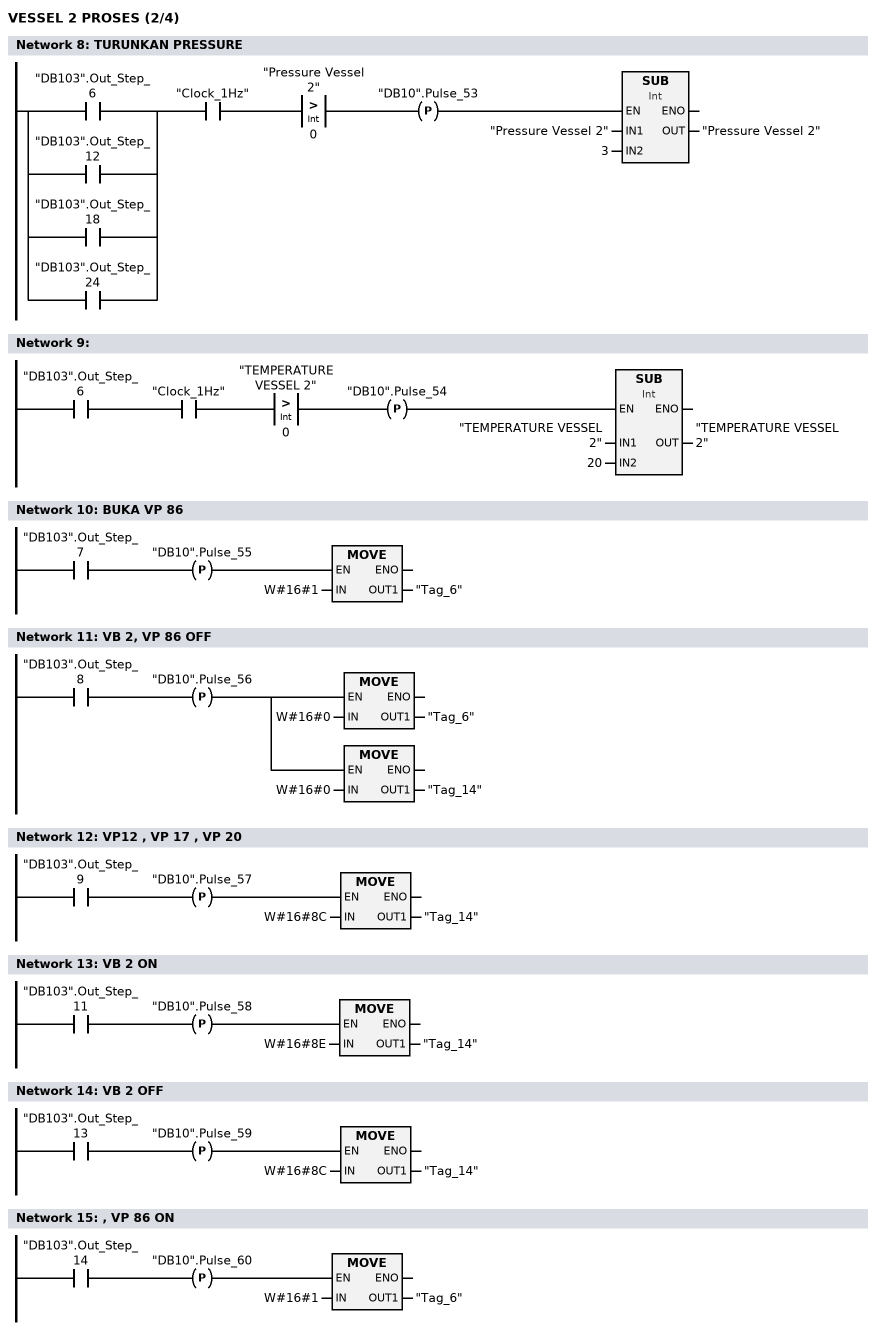
   RUNG wire#powerrail
      Contact( "DB103".Out_Step_6 )
      wire#w1
      Contact( "Clock_1Hz" )
      { S7_Templates := "SrcType := Int" } GT_Contact(in1 := "Pressure Vessel 2", in2 := 0)
      P_Trig( "DB10".Pulse_53 )
      { S7_Templates := "SrcType := Int" } Sub(in1 := "Pressure Vessel 2", in2 := 3, out => "Pressure Vessel 2")
   END_RUNG
   RUNG wire#powerrail
      Contact( "DB103".Out_Step_12 )
   END_RUNG wire#w1
   RUNG wire#powerrail
      Contact( "DB103".Out_Step_18 )
   END_RUNG wire#w1
   RUNG wire#powerrail
      Contact( "DB103".Out_Step_24 )
   END_RUNG wire#w1
   // the same network as SCL:
   #_w1 := ("DB103".Out_Step_6 OR "DB103".Out_Step_12 OR "DB103".Out_Step_18 OR "DB103".Out_Step_24) AND "Clock_1Hz" AND ("Pressure Vessel 2" > 0);
   #_w2 := #_w1 AND NOT "DB10".Pulse_53;   // rising edge
   "DB10".Pulse_53 := #_w1;
   IF #_w2 THEN "Pressure Vessel 2" := "Pressure Vessel 2" - 3; END_IF;
END_REGION

REGION Network 9
   RUNG wire#powerrail
      Contact( "DB103".Out_Step_6 )
      Contact( "Clock_1Hz" )
      { S7_Templates := "SrcType := Int" } GT_Contact(in1 := "TEMPERATURE VESSEL 2", in2 := 0)
      P_Trig( "DB10".Pulse_54 )
      { S7_Templates := "SrcType := Int" } Sub(in1 := "TEMPERATURE VESSEL 2", in2 := 20, out => "TEMPERATURE VESSEL 2")
   END_RUNG
   // the same network as SCL:
   #_w1 := "DB103".Out_Step_6 AND "Clock_1Hz" AND ("TEMPERATURE VESSEL 2" > 0);
   #_w2 := #_w1 AND NOT "DB10".Pulse_54;   // rising edge
   "DB10".Pulse_54 := #_w1;
   IF #_w2 THEN "TEMPERATURE VESSEL 2" := "TEMPERATURE VESSEL 2" - 20; END_IF;
END_REGION

REGION Network 10: BUKA VP 86
   RUNG wire#powerrail
      Contact( "DB103".Out_Step_7 )
      P_Trig( "DB10".Pulse_55 )
      Move(in := W#16#1, out1 => "Tag_6")
   END_RUNG
   // the same network as SCL:
   #_w1 := "DB103".Out_Step_7 AND NOT "DB10".Pulse_55;   // rising edge
   "DB10".Pulse_55 := "DB103".Out_Step_7;
   IF #_w1 THEN "Tag_6" := W#16#1; END_IF;
END_REGION

REGION Network 11: VB 2, VP 86 OFF
   RUNG wire#powerrail
      Contact( "DB103".Out_Step_8 )
      P_Trig( "DB10".Pulse_56 )
      wire#w1
      Move(in := W#16#0, out1 => "Tag_6")
   END_RUNG
   RUNG wire#w1
      Move(in := W#16#0, out1 => "Tag_14")
   END_RUNG
   // the same network as SCL:
   #_w1 := "DB103".Out_Step_8 AND NOT "DB10".Pulse_56;   // rising edge
   "DB10".Pulse_56 := "DB103".Out_Step_8;
   IF #_w1 THEN
       "Tag_6" := W#16#0;
       "Tag_14" := W#16#0;
   END_IF;
END_REGION

REGION Network 12: VP12 , VP 17 , VP 20
   RUNG wire#powerrail
      Contact( "DB103".Out_Step_9 )
      P_Trig( "DB10".Pulse_57 )
      Move(in := W#16#8C, out1 => "Tag_14")
   END_RUNG
   // the same network as SCL:
   #_w1 := "DB103".Out_Step_9 AND NOT "DB10".Pulse_57;   // rising edge
   "DB10".Pulse_57 := "DB103".Out_Step_9;
   IF #_w1 THEN "Tag_14" := W#16#8C; END_IF;
END_REGION

REGION Network 13: VB 2 ON
   RUNG wire#powerrail
      Contact( "DB103".Out_Step_11 )
      P_Trig( "DB10".Pulse_58 )
      Move(in := W#16#8E, out1 => "Tag_14")
   END_RUNG
   // the same network as SCL:
   #_w1 := "DB103".Out_Step_11 AND NOT "DB10".Pulse_58;   // rising edge
   "DB10".Pulse_58 := "DB103".Out_Step_11;
   IF #_w1 THEN "Tag_14" := W#16#8E; END_IF;
END_REGION

REGION Network 14: VB 2 OFF
   RUNG wire#powerrail
      Contact( "DB103".Out_Step_13 )
      P_Trig( "DB10".Pulse_59 )
      Move(in := W#16#8C, out1 => "Tag_14")
   END_RUNG
   // the same network as SCL:
   #_w1 := "DB103".Out_Step_13 AND NOT "DB10".Pulse_59;   // rising edge
   "DB10".Pulse_59 := "DB103".Out_Step_13;
   IF #_w1 THEN "Tag_14" := W#16#8C; END_IF;
END_REGION

REGION Network 15: , VP 86 ON
   RUNG wire#powerrail
      Contact( "DB103".Out_Step_14 )
      P_Trig( "DB10".Pulse_60 )
      Move(in := W#16#1, out1 => "Tag_6")
   END_RUNG
   // the same network as SCL:
   #_w1 := "DB103".Out_Step_14 AND NOT "DB10".Pulse_60;   // rising edge
   "DB10".Pulse_60 := "DB103".Out_Step_14;
   IF #_w1 THEN "Tag_6" := W#16#1; END_IF;
END_REGION

REGION Network 16: VP 86 OFF
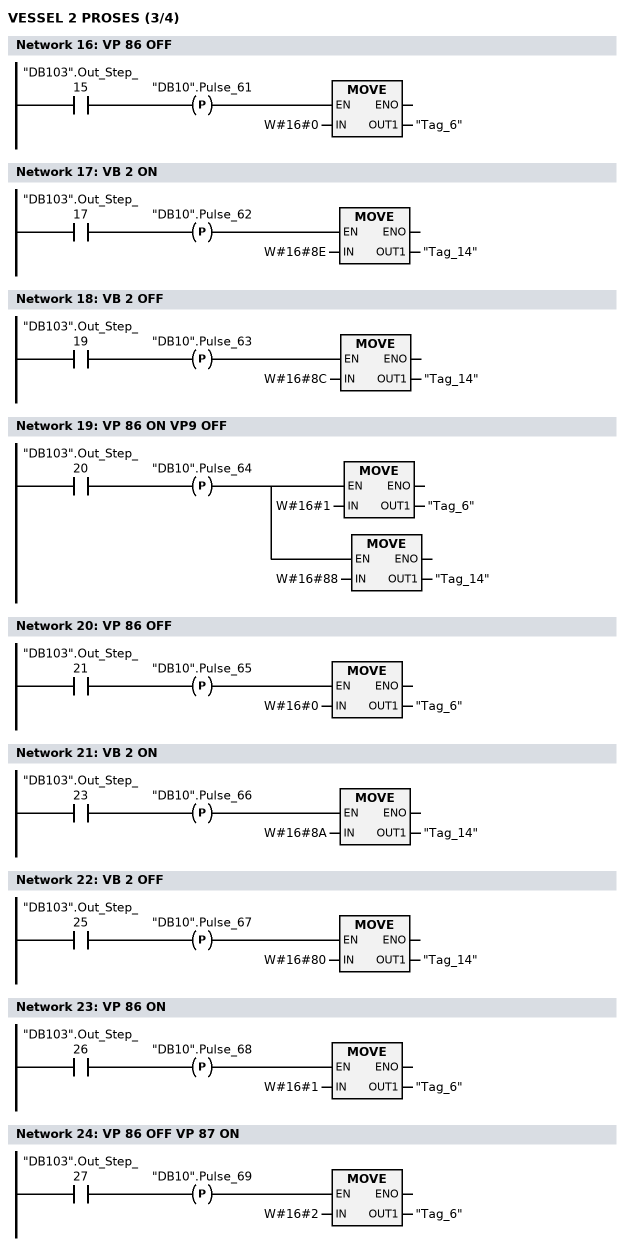
   RUNG wire#powerrail
      Contact( "DB103".Out_Step_15 )
      P_Trig( "DB10".Pulse_61 )
      Move(in := W#16#0, out1 => "Tag_6")
   END_RUNG
   // the same network as SCL:
   #_w1 := "DB103".Out_Step_15 AND NOT "DB10".Pulse_61;   // rising edge
   "DB10".Pulse_61 := "DB103".Out_Step_15;
   IF #_w1 THEN "Tag_6" := W#16#0; END_IF;
END_REGION

REGION Network 17: VB 2 ON
   RUNG wire#powerrail
      Contact( "DB103".Out_Step_17 )
      P_Trig( "DB10".Pulse_62 )
      Move(in := W#16#8E, out1 => "Tag_14")
   END_RUNG
   // the same network as SCL:
   #_w1 := "DB103".Out_Step_17 AND NOT "DB10".Pulse_62;   // rising edge
   "DB10".Pulse_62 := "DB103".Out_Step_17;
   IF #_w1 THEN "Tag_14" := W#16#8E; END_IF;
END_REGION

REGION Network 18: VB 2 OFF
   RUNG wire#powerrail
      Contact( "DB103".Out_Step_19 )
      P_Trig( "DB10".Pulse_63 )
      Move(in := W#16#8C, out1 => "Tag_14")
   END_RUNG
   // the same network as SCL:
   #_w1 := "DB103".Out_Step_19 AND NOT "DB10".Pulse_63;   // rising edge
   "DB10".Pulse_63 := "DB103".Out_Step_19;
   IF #_w1 THEN "Tag_14" := W#16#8C; END_IF;
END_REGION

REGION Network 19: VP 86 ON VP9 OFF
   RUNG wire#powerrail
      Contact( "DB103".Out_Step_20 )
      P_Trig( "DB10".Pulse_64 )
      wire#w1
      Move(in := W#16#1, out1 => "Tag_6")
   END_RUNG
   RUNG wire#w1
      Move(in := W#16#88, out1 => "Tag_14")
   END_RUNG
   // the same network as SCL:
   #_w1 := "DB103".Out_Step_20 AND NOT "DB10".Pulse_64;   // rising edge
   "DB10".Pulse_64 := "DB103".Out_Step_20;
   IF #_w1 THEN
       "Tag_6" := W#16#1;
       "Tag_14" := W#16#88;
   END_IF;
END_REGION

REGION Network 20: VP 86 OFF
   RUNG wire#powerrail
      Contact( "DB103".Out_Step_21 )
      P_Trig( "DB10".Pulse_65 )
      Move(in := W#16#0, out1 => "Tag_6")
   END_RUNG
   // the same network as SCL:
   #_w1 := "DB103".Out_Step_21 AND NOT "DB10".Pulse_65;   // rising edge
   "DB10".Pulse_65 := "DB103".Out_Step_21;
   IF #_w1 THEN "Tag_6" := W#16#0; END_IF;
END_REGION

REGION Network 21: VB 2 ON
   RUNG wire#powerrail
      Contact( "DB103".Out_Step_23 )
      P_Trig( "DB10".Pulse_66 )
      Move(in := W#16#8A, out1 => "Tag_14")
   END_RUNG
   // the same network as SCL:
   #_w1 := "DB103".Out_Step_23 AND NOT "DB10".Pulse_66;   // rising edge
   "DB10".Pulse_66 := "DB103".Out_Step_23;
   IF #_w1 THEN "Tag_14" := W#16#8A; END_IF;
END_REGION

REGION Network 22: VB 2 OFF
   RUNG wire#powerrail
      Contact( "DB103".Out_Step_25 )
      P_Trig( "DB10".Pulse_67 )
      Move(in := W#16#80, out1 => "Tag_14")
   END_RUNG
   // the same network as SCL:
   #_w1 := "DB103".Out_Step_25 AND NOT "DB10".Pulse_67;   // rising edge
   "DB10".Pulse_67 := "DB103".Out_Step_25;
   IF #_w1 THEN "Tag_14" := W#16#80; END_IF;
END_REGION

REGION Network 23: VP 86 ON
   RUNG wire#powerrail
      Contact( "DB103".Out_Step_26 )
      P_Trig( "DB10".Pulse_68 )
      Move(in := W#16#1, out1 => "Tag_6")
   END_RUNG
   // the same network as SCL:
   #_w1 := "DB103".Out_Step_26 AND NOT "DB10".Pulse_68;   // rising edge
   "DB10".Pulse_68 := "DB103".Out_Step_26;
   IF #_w1 THEN "Tag_6" := W#16#1; END_IF;
END_REGION

REGION Network 24: VP 86 OFF VP 87 ON
   RUNG wire#powerrail
      Contact( "DB103".Out_Step_27 )
      P_Trig( "DB10".Pulse_69 )
      Move(in := W#16#2, out1 => "Tag_6")
   END_RUNG
   // the same network as SCL:
   #_w1 := "DB103".Out_Step_27 AND NOT "DB10".Pulse_69;   // rising edge
   "DB10".Pulse_69 := "DB103".Out_Step_27;
   IF #_w1 THEN "Tag_6" := W#16#2; END_IF;
END_REGION

REGION Network 25: VP 87 OFF
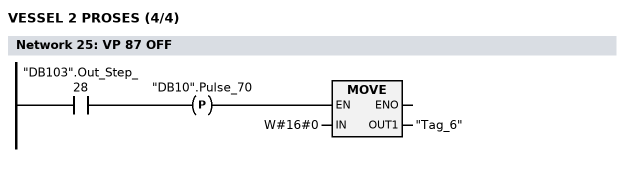
   RUNG wire#powerrail
      Contact( "DB103".Out_Step_28 )
      P_Trig( "DB10".Pulse_70 )
      Move(in := W#16#0, out1 => "Tag_6")
   END_RUNG
   // the same network as SCL:
   #_w1 := "DB103".Out_Step_28 AND NOT "DB10".Pulse_70;   // rising edge
   "DB10".Pulse_70 := "DB103".Out_Step_28;
   IF #_w1 THEN "Tag_6" := W#16#0; END_IF;
END_REGION
END_FUNCTION

FUNCTION "SEQUENCE V2 PROSES" : Void   // FC12, LAD
{ S7_Optimized_Access := 'TRUE' }
VERSION : 0.1
   VAR_TEMP   // added for the SCL form of the ladder/FBD networks
      _w1 : Bool;
      _w2 : Bool;
      _s5time1 : S5Time;
   END_VAR
BEGIN

REGION Network 1: START PROSES
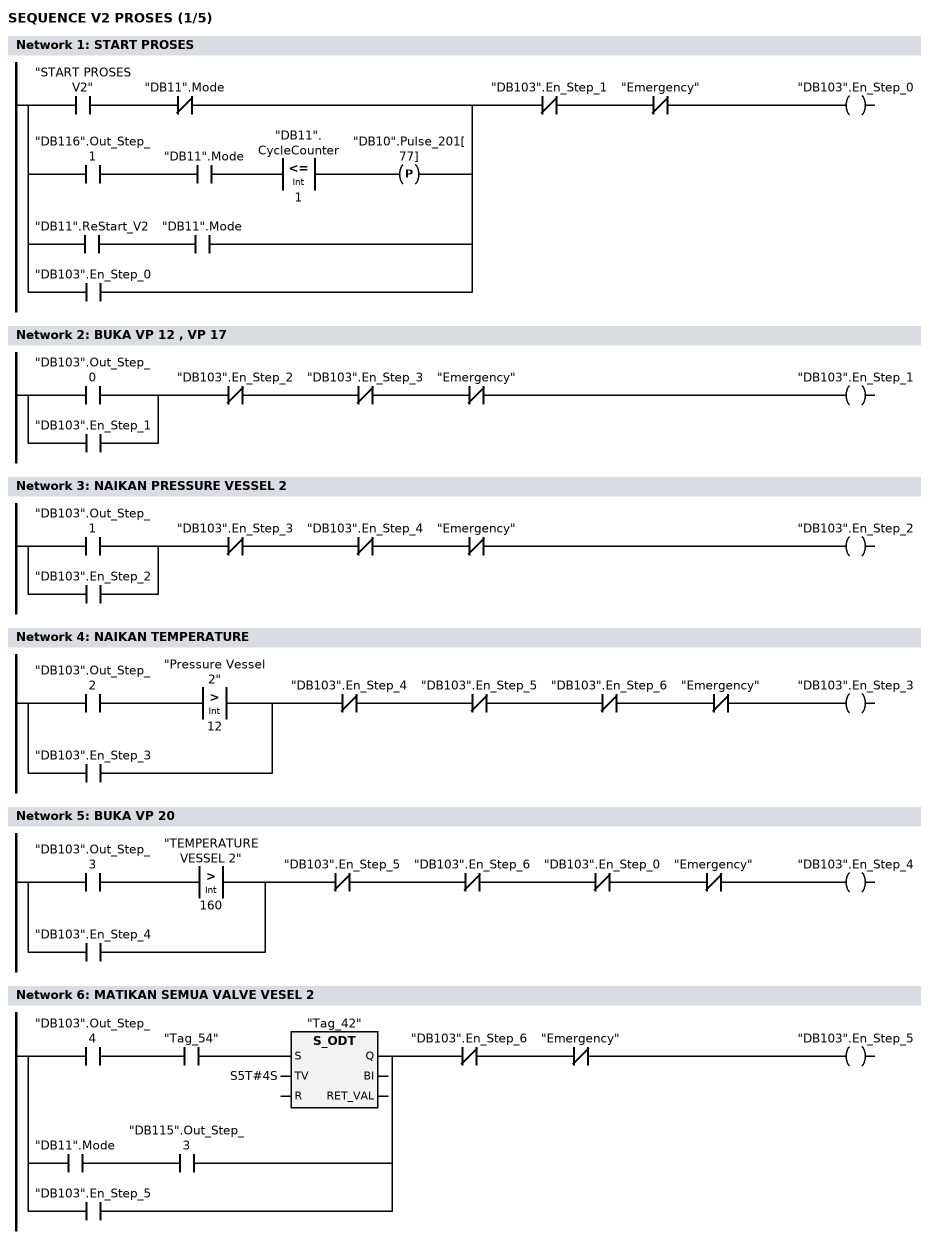
   RUNG wire#powerrail
      Contact( "START PROSES V2" )
      I_Contact( "DB11".Mode )
      wire#w1
      I_Contact( "DB103".En_Step_1 )
      I_Contact( "Emergency" )
      Coil( "DB103".En_Step_0 )
   END_RUNG
   RUNG wire#powerrail
      Contact( "DB116".Out_Step_1 )
      Contact( "DB11".Mode )
      { S7_Templates := "SrcType := Int" } LE_Contact(in1 := "DB11".CycleCounter, in2 := 1)
      P_Trig( "DB10".Pulse_201[77] )
   END_RUNG wire#w1
   RUNG wire#powerrail
      Contact( "DB11".ReStart_V2 )
      Contact( "DB11".Mode )
   END_RUNG wire#w1
   RUNG wire#powerrail
      Contact( "DB103".En_Step_0 )
   END_RUNG wire#w1
   // the same network as SCL:
   #_w1 := "DB116".Out_Step_1 AND "DB11".Mode AND ("DB11".CycleCounter <= 1);
   #_w2 := #_w1 AND NOT "DB10".Pulse_201[77];   // rising edge
   "DB10".Pulse_201[77] := #_w1;
   "DB103".En_Step_0 := (("START PROSES V2" AND NOT "DB11".Mode) OR #_w2 OR ("DB11".ReStart_V2 AND "DB11".Mode) OR "DB103".En_Step_0) AND NOT "DB103".En_Step_1 AND NOT "Emergency";
END_REGION

REGION Network 2: BUKA VP 12 , VP 17
   RUNG wire#powerrail
      Contact( "DB103".Out_Step_0 )
      wire#w1
      I_Contact( "DB103".En_Step_2 )
      I_Contact( "DB103".En_Step_3 )
      I_Contact( "Emergency" )
      Coil( "DB103".En_Step_1 )
   END_RUNG
   RUNG wire#powerrail
      Contact( "DB103".En_Step_1 )
   END_RUNG wire#w1
   // the same network as SCL:
   "DB103".En_Step_1 := ("DB103".Out_Step_0 OR "DB103".En_Step_1) AND NOT "DB103".En_Step_2 AND NOT "DB103".En_Step_3 AND NOT "Emergency";
END_REGION

REGION Network 3: NAIKAN PRESSURE VESSEL 2
   RUNG wire#powerrail
      Contact( "DB103".Out_Step_1 )
      wire#w1
      I_Contact( "DB103".En_Step_3 )
      I_Contact( "DB103".En_Step_4 )
      I_Contact( "Emergency" )
      Coil( "DB103".En_Step_2 )
   END_RUNG
   RUNG wire#powerrail
      Contact( "DB103".En_Step_2 )
   END_RUNG wire#w1
   // the same network as SCL:
   "DB103".En_Step_2 := ("DB103".Out_Step_1 OR "DB103".En_Step_2) AND NOT "DB103".En_Step_3 AND NOT "DB103".En_Step_4 AND NOT "Emergency";
END_REGION

REGION Network 4: NAIKAN TEMPERATURE
   RUNG wire#powerrail
      Contact( "DB103".Out_Step_2 )
      { S7_Templates := "SrcType := Int" } GT_Contact(in1 := "Pressure Vessel 2", in2 := 12)
      wire#w1
      I_Contact( "DB103".En_Step_4 )
      I_Contact( "DB103".En_Step_5 )
      I_Contact( "DB103".En_Step_6 )
      I_Contact( "Emergency" )
      Coil( "DB103".En_Step_3 )
   END_RUNG
   RUNG wire#powerrail
      Contact( "DB103".En_Step_3 )
   END_RUNG wire#w1
   // the same network as SCL:
   "DB103".En_Step_3 := (("DB103".Out_Step_2 AND ("Pressure Vessel 2" > 12)) OR "DB103".En_Step_3) AND NOT "DB103".En_Step_4 AND NOT "DB103".En_Step_5 AND NOT "DB103".En_Step_6 AND NOT "Emergency";
END_REGION

REGION Network 5: BUKA VP 20
   RUNG wire#powerrail
      Contact( "DB103".Out_Step_3 )
      { S7_Templates := "SrcType := Int" } GT_Contact(in1 := "TEMPERATURE VESSEL 2", in2 := 160)
      wire#w1
      I_Contact( "DB103".En_Step_5 )
      I_Contact( "DB103".En_Step_6 )
      I_Contact( "DB103".En_Step_0 )
      I_Contact( "Emergency" )
      Coil( "DB103".En_Step_4 )
   END_RUNG
   RUNG wire#powerrail
      Contact( "DB103".En_Step_4 )
   END_RUNG wire#w1
   // the same network as SCL:
   "DB103".En_Step_4 := (("DB103".Out_Step_3 AND ("TEMPERATURE VESSEL 2" > 160)) OR "DB103".En_Step_4) AND NOT "DB103".En_Step_5 AND NOT "DB103".En_Step_6 AND NOT "DB103".En_Step_0 AND NOT "Emergency";
END_REGION

REGION Network 6: MATIKAN SEMUA VALVE VESEL 2
   RUNG wire#powerrail
      Contact( "DB103".Out_Step_4 )
      Contact( "Tag_54" )
      S_ODT(T_NO := "Tag_42", TV := S5T#4S, R :=, BI =>, RET_VAL =>)
      wire#w1
      I_Contact( "DB103".En_Step_6 )
      I_Contact( "Emergency" )
      Coil( "DB103".En_Step_5 )
   END_RUNG
   RUNG wire#powerrail
      Contact( "DB11".Mode )
      Contact( "DB115".Out_Step_3 )
   END_RUNG wire#w1
   RUNG wire#powerrail
      Contact( "DB103".En_Step_5 )
   END_RUNG wire#w1
   // the same network as SCL:
   #_s5time1 := S_ODT(T_NO := "Tag_42", S := "DB103".Out_Step_4 AND "Tag_54", TV := S5T#4S, Q => #_w1);
   "DB103".En_Step_5 := (#_w1 OR ("DB11".Mode AND "DB115".Out_Step_3) OR "DB103".En_Step_5) AND NOT "DB103".En_Step_6 AND NOT "Emergency";
END_REGION

REGION Network 7: NYALAKAN VB 2
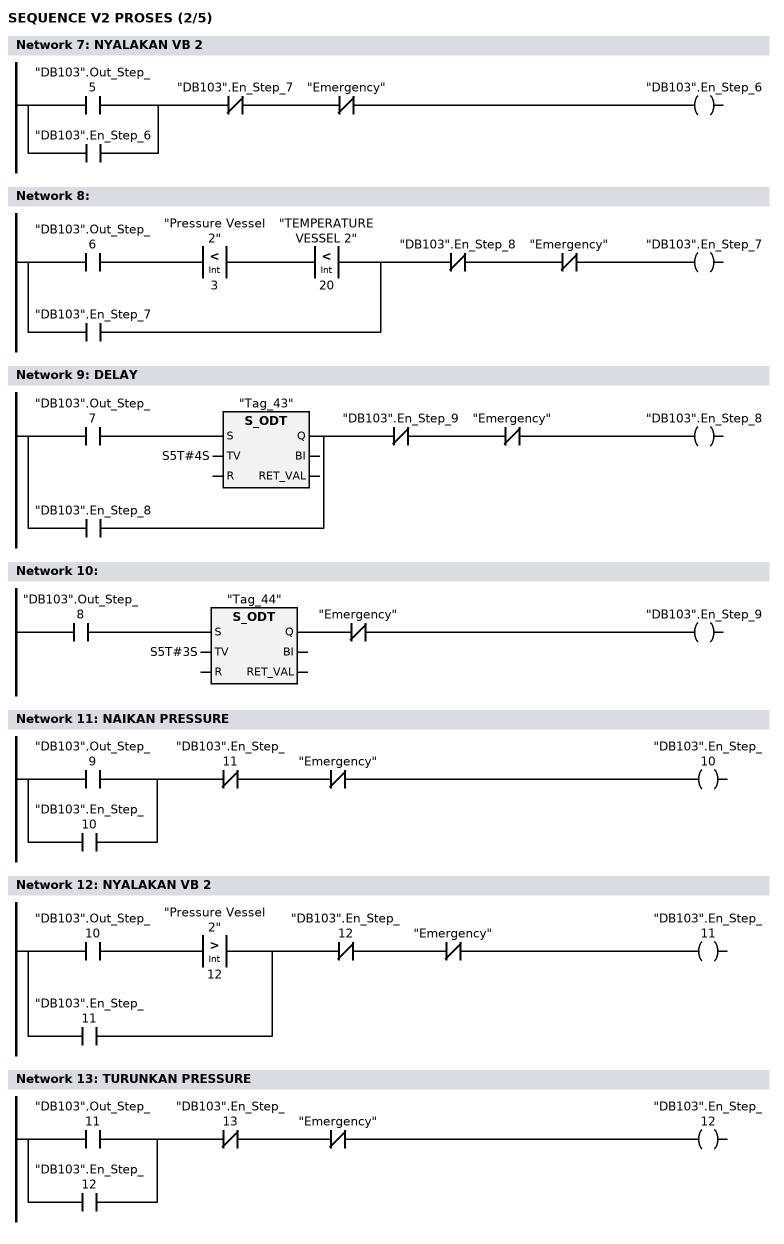
   RUNG wire#powerrail
      Contact( "DB103".Out_Step_5 )
      wire#w1
      I_Contact( "DB103".En_Step_7 )
      I_Contact( "Emergency" )
      Coil( "DB103".En_Step_6 )
   END_RUNG
   RUNG wire#powerrail
      Contact( "DB103".En_Step_6 )
   END_RUNG wire#w1
   // the same network as SCL:
   "DB103".En_Step_6 := ("DB103".Out_Step_5 OR "DB103".En_Step_6) AND NOT "DB103".En_Step_7 AND NOT "Emergency";
END_REGION

REGION Network 8
   RUNG wire#powerrail
      Contact( "DB103".Out_Step_6 )
      { S7_Templates := "SrcType := Int" } LT_Contact(in1 := "Pressure Vessel 2", in2 := 3)
      { S7_Templates := "SrcType := Int" } LT_Contact(in1 := "TEMPERATURE VESSEL 2", in2 := 20)
      wire#w1
      I_Contact( "DB103".En_Step_8 )
      I_Contact( "Emergency" )
      Coil( "DB103".En_Step_7 )
   END_RUNG
   RUNG wire#powerrail
      Contact( "DB103".En_Step_7 )
   END_RUNG wire#w1
   // the same network as SCL:
   "DB103".En_Step_7 := (("DB103".Out_Step_6 AND ("Pressure Vessel 2" < 3) AND ("TEMPERATURE VESSEL 2" < 20)) OR "DB103".En_Step_7) AND NOT "DB103".En_Step_8 AND NOT "Emergency";
END_REGION

REGION Network 9: DELAY
   RUNG wire#powerrail
      Contact( "DB103".Out_Step_7 )
      S_ODT(T_NO := "Tag_43", TV := S5T#4S, R :=, BI =>, RET_VAL =>)
      wire#w1
      I_Contact( "DB103".En_Step_9 )
      I_Contact( "Emergency" )
      Coil( "DB103".En_Step_8 )
   END_RUNG
   RUNG wire#powerrail
      Contact( "DB103".En_Step_8 )
   END_RUNG wire#w1
   // the same network as SCL:
   #_s5time1 := S_ODT(T_NO := "Tag_43", S := "DB103".Out_Step_7, TV := S5T#4S, Q => #_w1);
   "DB103".En_Step_8 := (#_w1 OR "DB103".En_Step_8) AND NOT "DB103".En_Step_9 AND NOT "Emergency";
END_REGION

REGION Network 10
   RUNG wire#powerrail
      Contact( "DB103".Out_Step_8 )
      S_ODT(T_NO := "Tag_44", TV := S5T#3S, R :=, BI =>, RET_VAL =>)
      I_Contact( "Emergency" )
      Coil( "DB103".En_Step_9 )
   END_RUNG
   // the same network as SCL:
   #_s5time1 := S_ODT(T_NO := "Tag_44", S := "DB103".Out_Step_8, TV := S5T#3S, Q => #_w1);
   "DB103".En_Step_9 := #_w1 AND NOT "Emergency";
END_REGION

REGION Network 11: NAIKAN PRESSURE
   RUNG wire#powerrail
      Contact( "DB103".Out_Step_9 )
      wire#w1
      I_Contact( "DB103".En_Step_11 )
      I_Contact( "Emergency" )
      Coil( "DB103".En_Step_10 )
   END_RUNG
   RUNG wire#powerrail
      Contact( "DB103".En_Step_10 )
   END_RUNG wire#w1
   // the same network as SCL:
   "DB103".En_Step_10 := ("DB103".Out_Step_9 OR "DB103".En_Step_10) AND NOT "DB103".En_Step_11 AND NOT "Emergency";
END_REGION

REGION Network 12: NYALAKAN VB 2
   RUNG wire#powerrail
      Contact( "DB103".Out_Step_10 )
      { S7_Templates := "SrcType := Int" } GT_Contact(in1 := "Pressure Vessel 2", in2 := 12)
      wire#w1
      I_Contact( "DB103".En_Step_12 )
      I_Contact( "Emergency" )
      Coil( "DB103".En_Step_11 )
   END_RUNG
   RUNG wire#powerrail
      Contact( "DB103".En_Step_11 )
   END_RUNG wire#w1
   // the same network as SCL:
   "DB103".En_Step_11 := (("DB103".Out_Step_10 AND ("Pressure Vessel 2" > 12)) OR "DB103".En_Step_11) AND NOT "DB103".En_Step_12 AND NOT "Emergency";
END_REGION

REGION Network 13: TURUNKAN PRESSURE
   RUNG wire#powerrail
      Contact( "DB103".Out_Step_11 )
      wire#w1
      I_Contact( "DB103".En_Step_13 )
      I_Contact( "Emergency" )
      Coil( "DB103".En_Step_12 )
   END_RUNG
   RUNG wire#powerrail
      Contact( "DB103".En_Step_12 )
   END_RUNG wire#w1
   // the same network as SCL:
   "DB103".En_Step_12 := ("DB103".Out_Step_11 OR "DB103".En_Step_12) AND NOT "DB103".En_Step_13 AND NOT "Emergency";
END_REGION

REGION Network 14
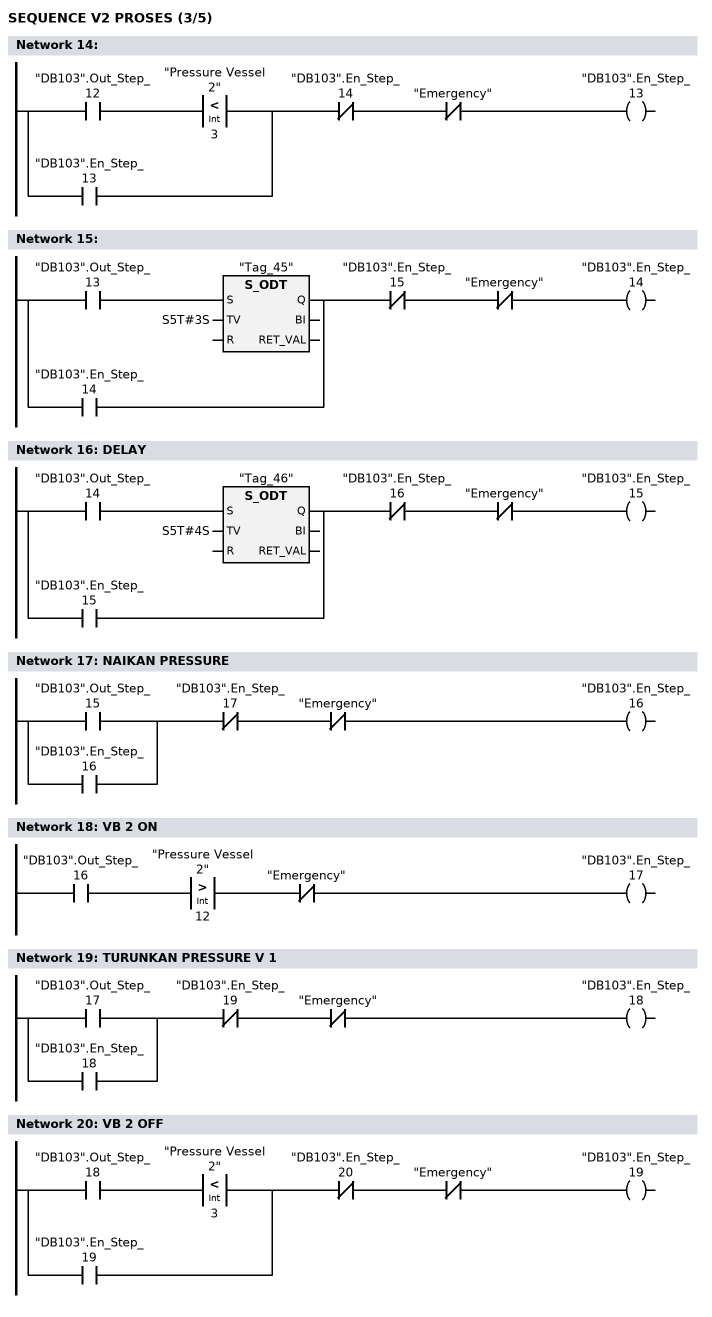
   RUNG wire#powerrail
      Contact( "DB103".Out_Step_12 )
      { S7_Templates := "SrcType := Int" } LT_Contact(in1 := "Pressure Vessel 2", in2 := 3)
      wire#w1
      I_Contact( "DB103".En_Step_14 )
      I_Contact( "Emergency" )
      Coil( "DB103".En_Step_13 )
   END_RUNG
   RUNG wire#powerrail
      Contact( "DB103".En_Step_13 )
   END_RUNG wire#w1
   // the same network as SCL:
   "DB103".En_Step_13 := (("DB103".Out_Step_12 AND ("Pressure Vessel 2" < 3)) OR "DB103".En_Step_13) AND NOT "DB103".En_Step_14 AND NOT "Emergency";
END_REGION

REGION Network 15
   RUNG wire#powerrail
      Contact( "DB103".Out_Step_13 )
      S_ODT(T_NO := "Tag_45", TV := S5T#3S, R :=, BI =>, RET_VAL =>)
      wire#w1
      I_Contact( "DB103".En_Step_15 )
      I_Contact( "Emergency" )
      Coil( "DB103".En_Step_14 )
   END_RUNG
   RUNG wire#powerrail
      Contact( "DB103".En_Step_14 )
   END_RUNG wire#w1
   // the same network as SCL:
   #_s5time1 := S_ODT(T_NO := "Tag_45", S := "DB103".Out_Step_13, TV := S5T#3S, Q => #_w1);
   "DB103".En_Step_14 := (#_w1 OR "DB103".En_Step_14) AND NOT "DB103".En_Step_15 AND NOT "Emergency";
END_REGION

REGION Network 16: DELAY
   RUNG wire#powerrail
      Contact( "DB103".Out_Step_14 )
      S_ODT(T_NO := "Tag_46", TV := S5T#4S, R :=, BI =>, RET_VAL =>)
      wire#w1
      I_Contact( "DB103".En_Step_16 )
      I_Contact( "Emergency" )
      Coil( "DB103".En_Step_15 )
   END_RUNG
   RUNG wire#powerrail
      Contact( "DB103".En_Step_15 )
   END_RUNG wire#w1
   // the same network as SCL:
   #_s5time1 := S_ODT(T_NO := "Tag_46", S := "DB103".Out_Step_14, TV := S5T#4S, Q => #_w1);
   "DB103".En_Step_15 := (#_w1 OR "DB103".En_Step_15) AND NOT "DB103".En_Step_16 AND NOT "Emergency";
END_REGION

REGION Network 17: NAIKAN PRESSURE
   RUNG wire#powerrail
      Contact( "DB103".Out_Step_15 )
      wire#w1
      I_Contact( "DB103".En_Step_17 )
      I_Contact( "Emergency" )
      Coil( "DB103".En_Step_16 )
   END_RUNG
   RUNG wire#powerrail
      Contact( "DB103".En_Step_16 )
   END_RUNG wire#w1
   // the same network as SCL:
   "DB103".En_Step_16 := ("DB103".Out_Step_15 OR "DB103".En_Step_16) AND NOT "DB103".En_Step_17 AND NOT "Emergency";
END_REGION

REGION Network 18: VB 2 ON
   RUNG wire#powerrail
      Contact( "DB103".Out_Step_16 )
      { S7_Templates := "SrcType := Int" } GT_Contact(in1 := "Pressure Vessel 2", in2 := 12)
      I_Contact( "Emergency" )
      Coil( "DB103".En_Step_17 )
   END_RUNG
   // the same network as SCL:
   "DB103".En_Step_17 := "DB103".Out_Step_16 AND ("Pressure Vessel 2" > 12) AND NOT "Emergency";
END_REGION

REGION Network 19: TURUNKAN PRESSURE V 1
   RUNG wire#powerrail
      Contact( "DB103".Out_Step_17 )
      wire#w1
      I_Contact( "DB103".En_Step_19 )
      I_Contact( "Emergency" )
      Coil( "DB103".En_Step_18 )
   END_RUNG
   RUNG wire#powerrail
      Contact( "DB103".En_Step_18 )
   END_RUNG wire#w1
   // the same network as SCL:
   "DB103".En_Step_18 := ("DB103".Out_Step_17 OR "DB103".En_Step_18) AND NOT "DB103".En_Step_19 AND NOT "Emergency";
END_REGION

REGION Network 20: VB 2 OFF
   RUNG wire#powerrail
      Contact( "DB103".Out_Step_18 )
      { S7_Templates := "SrcType := Int" } LT_Contact(in1 := "Pressure Vessel 2", in2 := 3)
      wire#w1
      I_Contact( "DB103".En_Step_20 )
      I_Contact( "Emergency" )
      Coil( "DB103".En_Step_19 )
   END_RUNG
   RUNG wire#powerrail
      Contact( "DB103".En_Step_19 )
   END_RUNG wire#w1
   // the same network as SCL:
   "DB103".En_Step_19 := (("DB103".Out_Step_18 AND ("Pressure Vessel 2" < 3)) OR "DB103".En_Step_19) AND NOT "DB103".En_Step_20 AND NOT "Emergency";
END_REGION

REGION Network 21: VP 86 ON VP 1 OFF
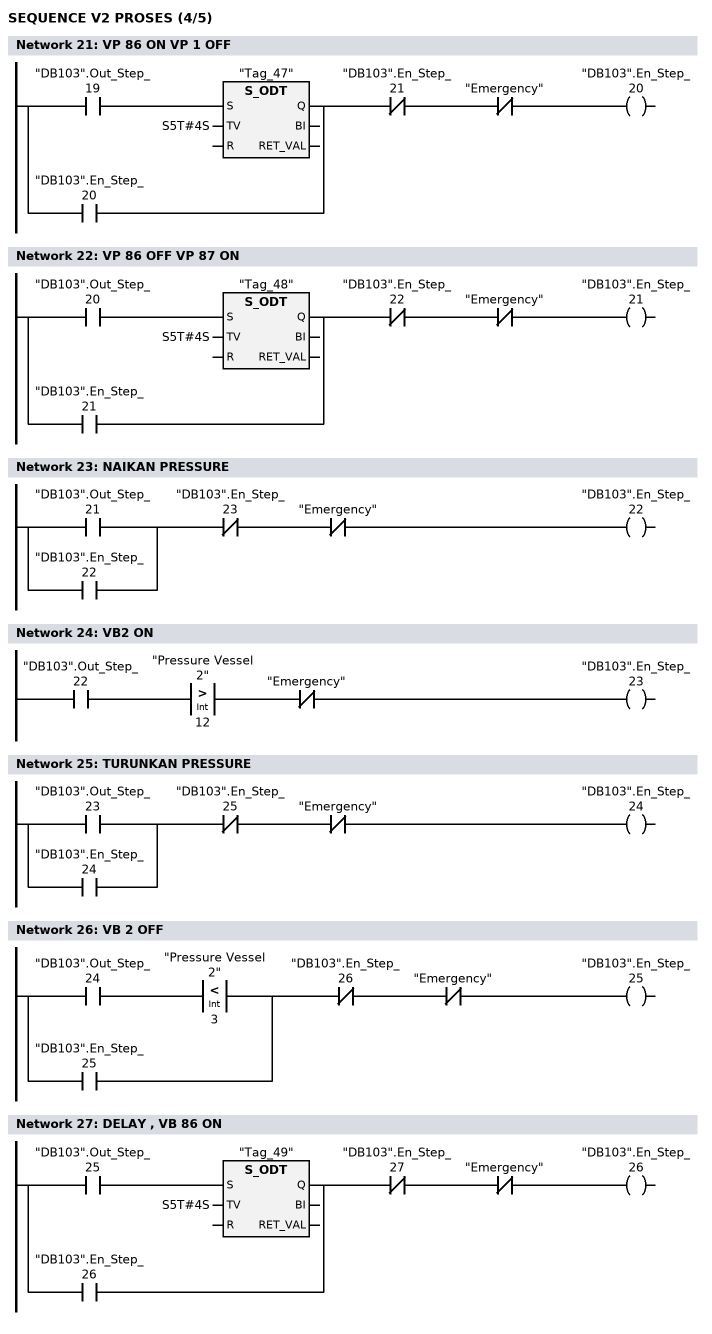
   RUNG wire#powerrail
      Contact( "DB103".Out_Step_19 )
      S_ODT(T_NO := "Tag_47", TV := S5T#4S, R :=, BI =>, RET_VAL =>)
      wire#w1
      I_Contact( "DB103".En_Step_21 )
      I_Contact( "Emergency" )
      Coil( "DB103".En_Step_20 )
   END_RUNG
   RUNG wire#powerrail
      Contact( "DB103".En_Step_20 )
   END_RUNG wire#w1
   // the same network as SCL:
   #_s5time1 := S_ODT(T_NO := "Tag_47", S := "DB103".Out_Step_19, TV := S5T#4S, Q => #_w1);
   "DB103".En_Step_20 := (#_w1 OR "DB103".En_Step_20) AND NOT "DB103".En_Step_21 AND NOT "Emergency";
END_REGION

REGION Network 22: VP 86 OFF VP 87 ON
   RUNG wire#powerrail
      Contact( "DB103".Out_Step_20 )
      S_ODT(T_NO := "Tag_48", TV := S5T#4S, R :=, BI =>, RET_VAL =>)
      wire#w1
      I_Contact( "DB103".En_Step_22 )
      I_Contact( "Emergency" )
      Coil( "DB103".En_Step_21 )
   END_RUNG
   RUNG wire#powerrail
      Contact( "DB103".En_Step_21 )
   END_RUNG wire#w1
   // the same network as SCL:
   #_s5time1 := S_ODT(T_NO := "Tag_48", S := "DB103".Out_Step_20, TV := S5T#4S, Q => #_w1);
   "DB103".En_Step_21 := (#_w1 OR "DB103".En_Step_21) AND NOT "DB103".En_Step_22 AND NOT "Emergency";
END_REGION

REGION Network 23: NAIKAN PRESSURE
   RUNG wire#powerrail
      Contact( "DB103".Out_Step_21 )
      wire#w1
      I_Contact( "DB103".En_Step_23 )
      I_Contact( "Emergency" )
      Coil( "DB103".En_Step_22 )
   END_RUNG
   RUNG wire#powerrail
      Contact( "DB103".En_Step_22 )
   END_RUNG wire#w1
   // the same network as SCL:
   "DB103".En_Step_22 := ("DB103".Out_Step_21 OR "DB103".En_Step_22) AND NOT "DB103".En_Step_23 AND NOT "Emergency";
END_REGION

REGION Network 24: VB2 ON
   RUNG wire#powerrail
      Contact( "DB103".Out_Step_22 )
      { S7_Templates := "SrcType := Int" } GT_Contact(in1 := "Pressure Vessel 2", in2 := 12)
      I_Contact( "Emergency" )
      Coil( "DB103".En_Step_23 )
   END_RUNG
   // the same network as SCL:
   "DB103".En_Step_23 := "DB103".Out_Step_22 AND ("Pressure Vessel 2" > 12) AND NOT "Emergency";
END_REGION

REGION Network 25: TURUNKAN PRESSURE
   RUNG wire#powerrail
      Contact( "DB103".Out_Step_23 )
      wire#w1
      I_Contact( "DB103".En_Step_25 )
      I_Contact( "Emergency" )
      Coil( "DB103".En_Step_24 )
   END_RUNG
   RUNG wire#powerrail
      Contact( "DB103".En_Step_24 )
   END_RUNG wire#w1
   // the same network as SCL:
   "DB103".En_Step_24 := ("DB103".Out_Step_23 OR "DB103".En_Step_24) AND NOT "DB103".En_Step_25 AND NOT "Emergency";
END_REGION

REGION Network 26: VB 2 OFF
   RUNG wire#powerrail
      Contact( "DB103".Out_Step_24 )
      { S7_Templates := "SrcType := Int" } LT_Contact(in1 := "Pressure Vessel 2", in2 := 3)
      wire#w1
      I_Contact( "DB103".En_Step_26 )
      I_Contact( "Emergency" )
      Coil( "DB103".En_Step_25 )
   END_RUNG
   RUNG wire#powerrail
      Contact( "DB103".En_Step_25 )
   END_RUNG wire#w1
   // the same network as SCL:
   "DB103".En_Step_25 := (("DB103".Out_Step_24 AND ("Pressure Vessel 2" < 3)) OR "DB103".En_Step_25) AND NOT "DB103".En_Step_26 AND NOT "Emergency";
END_REGION

REGION Network 27: DELAY , VB 86 ON
   RUNG wire#powerrail
      Contact( "DB103".Out_Step_25 )
      S_ODT(T_NO := "Tag_49", TV := S5T#4S, R :=, BI =>, RET_VAL =>)
      wire#w1
      I_Contact( "DB103".En_Step_27 )
      I_Contact( "Emergency" )
      Coil( "DB103".En_Step_26 )
   END_RUNG
   RUNG wire#powerrail
      Contact( "DB103".En_Step_26 )
   END_RUNG wire#w1
   // the same network as SCL:
   #_s5time1 := S_ODT(T_NO := "Tag_49", S := "DB103".Out_Step_25, TV := S5T#4S, Q => #_w1);
   "DB103".En_Step_26 := (#_w1 OR "DB103".En_Step_26) AND NOT "DB103".En_Step_27 AND NOT "Emergency";
END_REGION

REGION Network 28: VB 86 OFF VB 87 ON
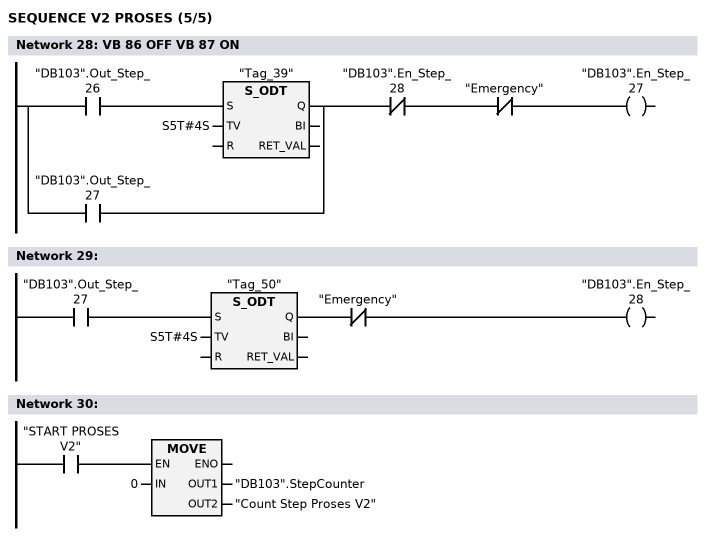
   RUNG wire#powerrail
      Contact( "DB103".Out_Step_26 )
      S_ODT(T_NO := "Tag_39", TV := S5T#4S, R :=, BI =>, RET_VAL =>)
      wire#w1
      I_Contact( "DB103".En_Step_28 )
      I_Contact( "Emergency" )
      Coil( "DB103".En_Step_27 )
   END_RUNG
   RUNG wire#powerrail
      Contact( "DB103".Out_Step_27 )
   END_RUNG wire#w1
   // the same network as SCL:
   #_s5time1 := S_ODT(T_NO := "Tag_39", S := "DB103".Out_Step_26, TV := S5T#4S, Q => #_w1);
   "DB103".En_Step_27 := (#_w1 OR "DB103".Out_Step_27) AND NOT "DB103".En_Step_28 AND NOT "Emergency";
END_REGION

REGION Network 29
   RUNG wire#powerrail
      Contact( "DB103".Out_Step_27 )
      S_ODT(T_NO := "Tag_50", TV := S5T#4S, R :=, BI =>, RET_VAL =>)
      I_Contact( "Emergency" )
      Coil( "DB103".En_Step_28 )
   END_RUNG
   // the same network as SCL:
   #_s5time1 := S_ODT(T_NO := "Tag_50", S := "DB103".Out_Step_27, TV := S5T#4S, Q => #_w1);
   "DB103".En_Step_28 := #_w1 AND NOT "Emergency";
END_REGION

REGION Network 30
   RUNG wire#powerrail
      Contact( "START PROSES V2" )
      Move(in := 0, out1 => "DB103".StepCounter, out2 => "Count Step Proses V2")
   END_RUNG
   // the same network as SCL:
   IF "START PROSES V2" THEN
       "DB103".StepCounter := 0;
       "Count Step Proses V2" := 0;
   END_IF;
END_REGION
END_FUNCTION

FUNCTION "VESSEL 3 PROSES" : Void   // FC13, LAD
{ S7_Optimized_Access := 'TRUE' }
VERSION : 0.1
   VAR_TEMP   // added for the SCL form of the ladder/FBD networks
      _w1 : Bool;
      _w2 : Bool;
   END_VAR
BEGIN

REGION Network 1: BUKA VALVE VP 12 DAN VP 17
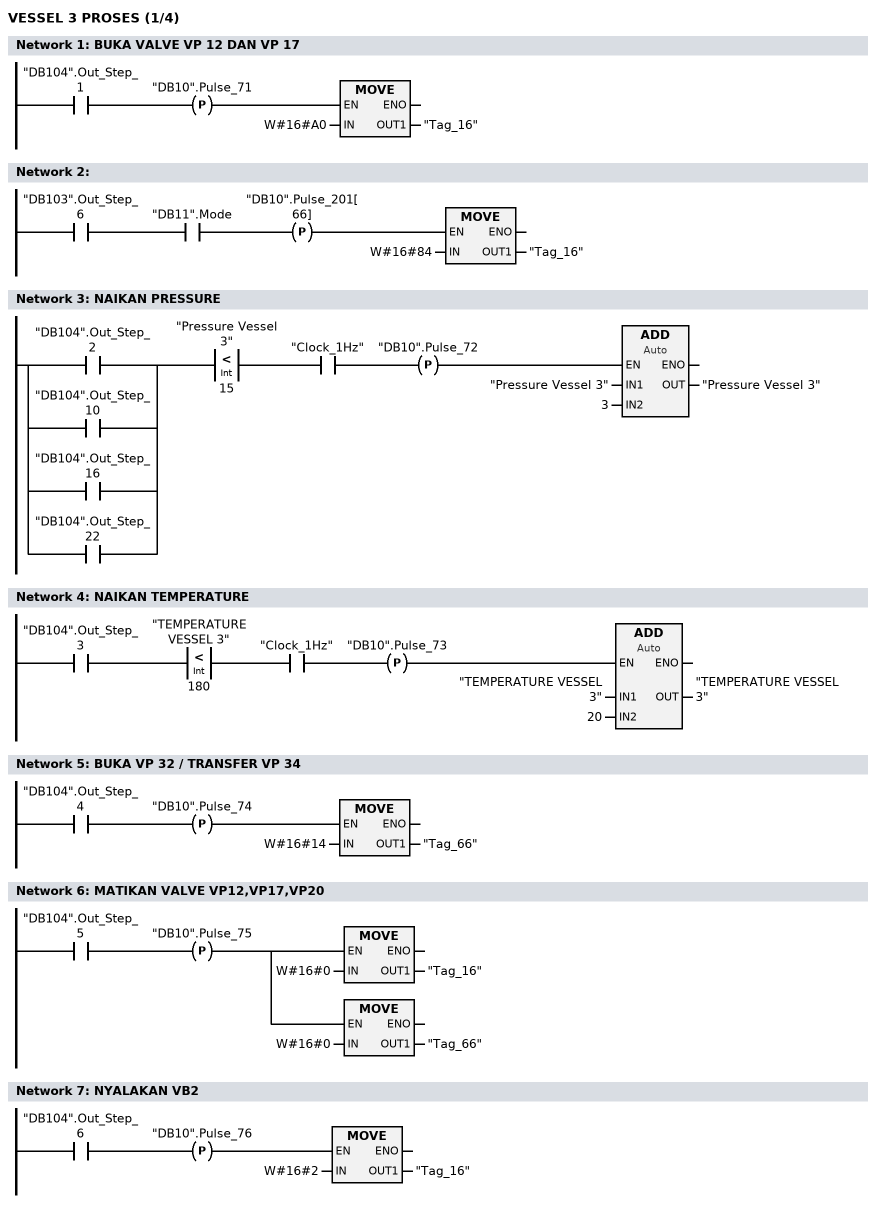
   RUNG wire#powerrail
      Contact( "DB104".Out_Step_1 )
      P_Trig( "DB10".Pulse_71 )
      Move(in := W#16#A0, out1 => "Tag_16")
   END_RUNG
   // the same network as SCL:
   #_w1 := "DB104".Out_Step_1 AND NOT "DB10".Pulse_71;   // rising edge
   "DB10".Pulse_71 := "DB104".Out_Step_1;
   IF #_w1 THEN "Tag_16" := W#16#A0; END_IF;
END_REGION
